(* Logix 5000 project; controller FV vendor 1 type 14 code 217 rev 31.11; software revision 31.00; part 44 of 63 *)
(* tags used below, declared in another part *)
   Dummy : BOOL;
   FV_B211 : DINT[255];   // GLYCL_SEL Glycol Pump Selectio n Words
   FV_B211_3_12_OutputBit : BOOL;
   FV_B211_3_13_OutputBit : BOOL;
   FV_B211_3_14_OutputBit : BOOL;
   fv_data_file_value_to_move : DINT;
   FV_from_data_file : DINT;
   FV_from_data_offset : DINT;
   FV_FV23C : PlantItem;   // FV23C
   FV_FV23J : PlantItem;   // FV23J
   FV_FV24C : PlantItem;   // FV24C
   FV_FV24J : PlantItem;   // FV24J
   FV_FV25C : PlantItem;   // FV25C
   FV_FV25J : PlantItem;   // FV25J
   FV_FV26C : PlantItem;   // FV26C
   FV_FV26J : PlantItem;   // FV26J
   FV_FV27C : PlantItem;   // FV27C
   FV_FV27J : PlantItem;   // FV27J
   FV_FV28C : PlantItem;   // FV28C
   FV_FV28J : PlantItem;   // FV28J
   FV_FV29C : PlantItem;   // FV29C
   FV_FV29J : PlantItem;   // FV29J
   FV_FV30C : PlantItem;   // FV30C
   FV_FV30J : PlantItem;   // FV30J
   FV_FV31C : PlantItem;   // FV31C
   FV_FV31J : PlantItem;   // FV31J
   FV_N110 : INT[255];   // FV DATA 0 CURRENT FV DATA
   FV_N111 : INT[50];   // FV1, CURRENT FV DATA
   FV_N112 : INT[50];   // FV2, CURRENT FV DATA
   FV_N113 : INT[50];   // FV3, CURRENT FV DATA
   FV_N114 : INT[50];   // FV4, CURRENT FV DATA
   FV_N115 : INT[50];   // FV5, CURRENT FV DATA
   FV_N116 : INT[50];   // FV6, CURRENT FV DATA
   FV_N117 : INT[50];   // FV7, CURRENT FV DATA
   FV_N118 : INT[50];   // FV8, CURRENT FV DATA
   FV_N119 : INT[50];   // FV9, CURRENT FV DATA
   FV_N120 : INT[50];   // FV10, CURRENT FV DATA
   FV_N121 : INT[50];   // FV11, CURRENT FV DATA
   FV_N122 : INT[50];   // FV12, CURRENT FV DATA
   FV_N123 : INT[50];   // FV13, CURRENT FV DATA
   FV_N124 : INT[50];   // FV14, CURRENT FV DATA
   FV_N125 : INT[50];   // FV15, CURRENT FV DATA
   FV_N126 : INT[50];   // FV16, CURRENT FV DATA
   FV_N127 : INT[50];   // FV17, CURRENT FV DATA
   FV_N128 : INT[50];   // FV18, CURRENT FV DATA
   FV_N129 : INT[50];   // FV19, CURRENT FV DATA
   FV_N130 : INT[50];   // FV20, CURRENT FV DATA
   FV_N131 : INT[50];   // FV21, CURRENT FV DATA
   FV_N132 : INT[50];   // FV22, CURRENT FV DATA
   FV_N133 : INT[50];   // FV23, CURRENT FV DATA
   FV_N134 : INT[50];   // FV24, CURRENT FV DATA
   FV_N135 : INT[50];   // FV25, CURRENT FV DATA
   FV_N136 : INT[50];   // YSV1, CURRENT FV DATA
   FV_N137 : INT[50];   // YSV2, CURRENT FV DATA
   FV_N138 : INT[50];   // YSV3, CURRENT FV DATA
   FV_N139 : INT[255];   // YST1
   FV_N140 : INT[255];   // YST2
   FV_N141 : INT[255];   // YSV1 DATA
   FV_N142 : INT[255];   // YSV2 DATA
   FV_N143 : INT[255];   // YSV3 DATA
   FV_N144 : INT[255];   // YST1 DATA
   FV_N145 : INT[255];   // YST2 DATA
   FV_N146 : INT[50];   // FV26, CURRENT FV DATA
   FV_N147 : INT[50];   // FV27, CURRENT FV DATA
   FV_N148 : INT[50];   // FV28, CURRENT FV DATA
   FV_N149 : INT[50];   // FV29, CURRENT FV DATA
   FV_N150 : INT[50];   // FV30, CURRENT FV DATA
   FV_N151 : INT[50];   // FV31, CURRENT FV DATA
   FV_N210 : INT[255];   // GLYCL_PTRS
   FV_PUMP1 : PlantItem;   // PUMP1
   FV_PUMP2 : PlantItem;   // PUMP2
   FV_PUMP3 : PlantItem;   // PUMP3
   FV_R6 : CONTROL[5];
   FV_SFile : INT[255];   // SLC Equivalent System File, So Original Code Can Remain
   FV_T212 : TIMER[5];
   FV_YSV1CV : PlantItem;   // YSV1CV
   FV_YSV1J : PlantItem;   // YSV1J
   FV_YSV2CV : PlantItem;   // YSV2CV
   FV_YSV2J : PlantItem;   // YSV2J
   FV_YSV3J : PlantItem;   // YSV3J
   MV_YST_Levels : REAL[2];
   YP_AV2 : PlantItem;   // AV2
   YST_BL_PMP_ON : BOOL;   // Blunger Pump
(* FV_Common, continued *)

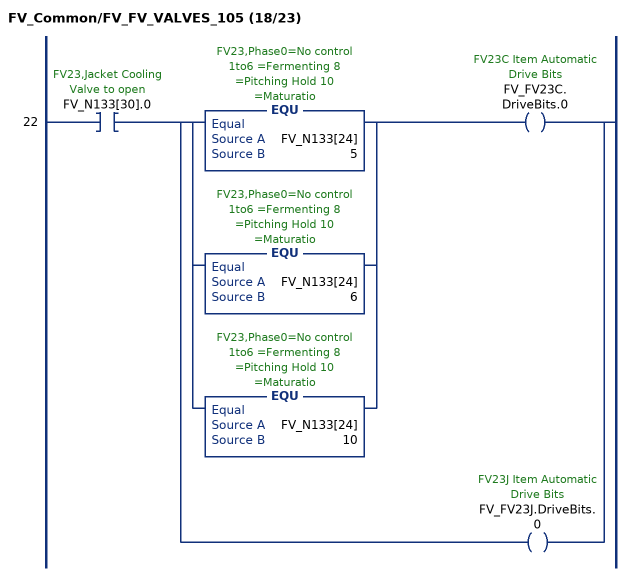
   [picture p944: FV_Common/FV_FV_VALVES_105 rungs 22-22]
   22: XIC(FV_N133[30].0)[[EQU(FV_N133[24],5) ,EQU(FV_N133[24],6) ,EQU(FV_N133[24],10) ] OTE(FV_FV23C.DriveBits.0) ,OTE(FV_FV23J.DriveBits.0) ];
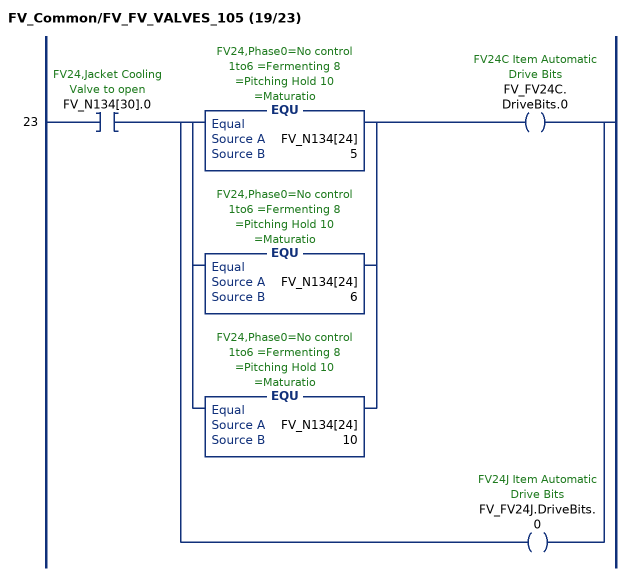
   23: XIC(FV_N134[30].0)[[EQU(FV_N134[24],5) ,EQU(FV_N134[24],6) ,EQU(FV_N134[24],10) ] OTE(FV_FV24C.DriveBits.0) ,OTE(FV_FV24J.DriveBits.0) ];
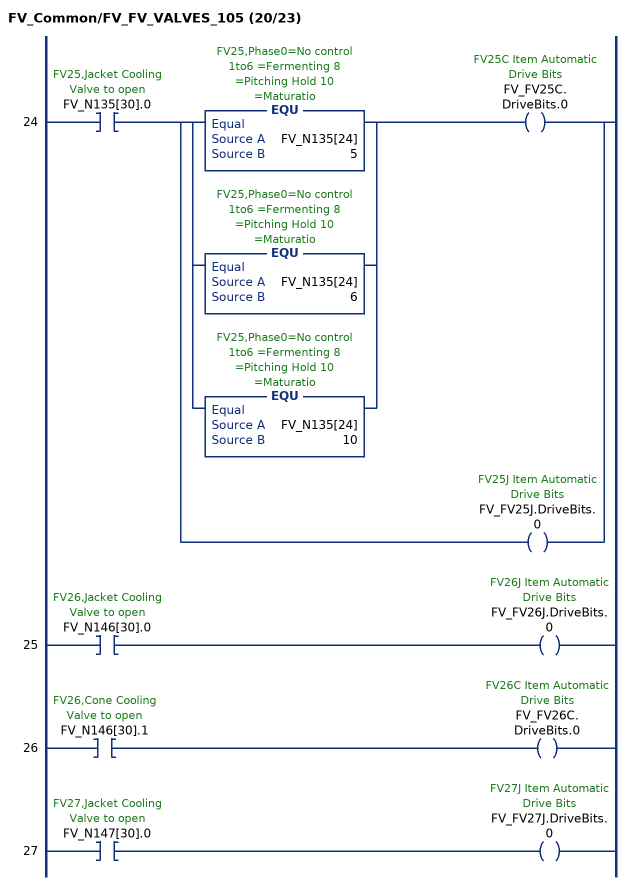
   24: XIC(FV_N135[30].0)[[EQU(FV_N135[24],5) ,EQU(FV_N135[24],6) ,EQU(FV_N135[24],10) ] OTE(FV_FV25C.DriveBits.0) ,OTE(FV_FV25J.DriveBits.0) ];
   25: XIC(FV_N146[30].0)OTE(FV_FV26J.DriveBits.0);
   26: XIC(FV_N146[30].1)OTE(FV_FV26C.DriveBits.0);
   27: XIC(FV_N147[30].0)OTE(FV_FV27J.DriveBits.0);
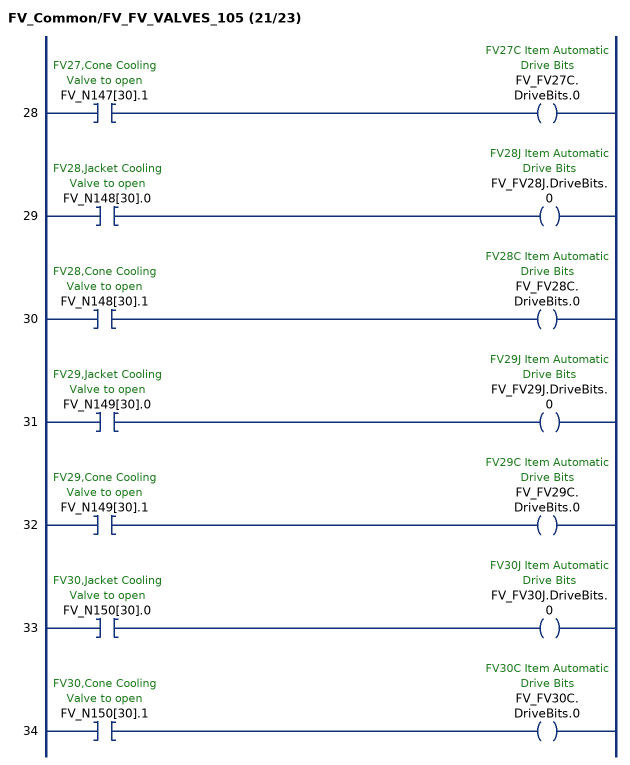
   28: XIC(FV_N147[30].1)OTE(FV_FV27C.DriveBits.0);
   29: XIC(FV_N148[30].0)OTE(FV_FV28J.DriveBits.0);
   30: XIC(FV_N148[30].1)OTE(FV_FV28C.DriveBits.0);
   31: XIC(FV_N149[30].0)OTE(FV_FV29J.DriveBits.0);
   32: XIC(FV_N149[30].1)OTE(FV_FV29C.DriveBits.0);
   33: XIC(FV_N150[30].0)OTE(FV_FV30J.DriveBits.0);
   34: XIC(FV_N150[30].1)OTE(FV_FV30C.DriveBits.0);
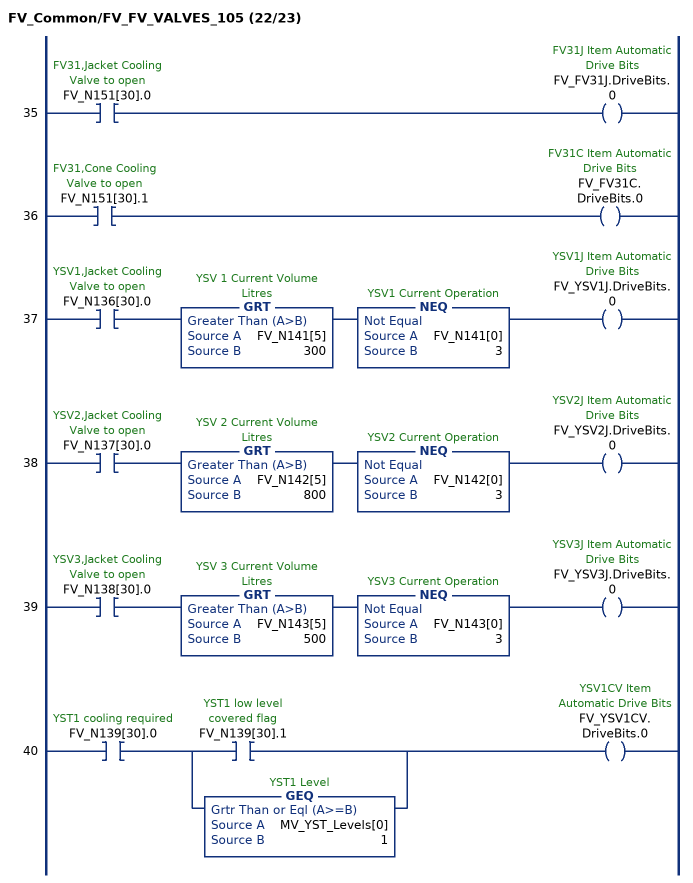
   35: XIC(FV_N151[30].0)OTE(FV_FV31J.DriveBits.0);
   36: XIC(FV_N151[30].1)OTE(FV_FV31C.DriveBits.0);
   37: XIC(FV_N136[30].0)GRT(FV_N141[5],300)NEQ(FV_N141[0],3)OTE(FV_YSV1J.DriveBits.0);
   38: XIC(FV_N137[30].0)GRT(FV_N142[5],800)NEQ(FV_N142[0],3)OTE(FV_YSV2J.DriveBits.0);
   39: XIC(FV_N138[30].0)GRT(FV_N143[5],500)NEQ(FV_N143[0],3)OTE(FV_YSV3J.DriveBits.0);
   40: XIC(FV_N139[30].0)[XIC(FV_N139[30].1) ,GEQ(MV_YST_Levels[0],1) ]OTE(FV_YSV1CV.DriveBits.0);
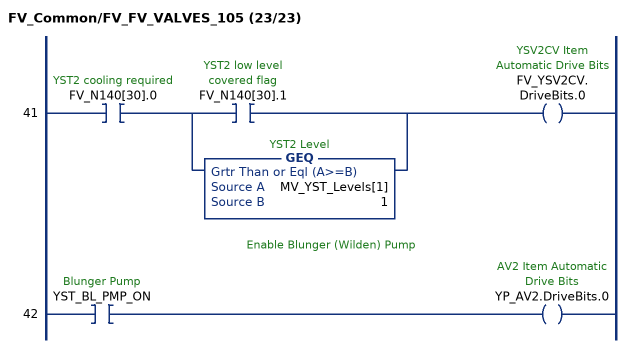
   41: XIC(FV_N140[30].0)[XIC(FV_N140[30].1) ,GEQ(MV_YST_Levels[1],1) ]OTE(FV_YSV2CV.DriveBits.0);
   // Enable Blunger (Wilden) Pump
   42: XIC(YST_BL_PMP_ON)OTE(YP_AV2.DriveBits.0);
END_ROUTINE

ROUTINE FV_Get_FV_Datafile_Value   (* ladder *)
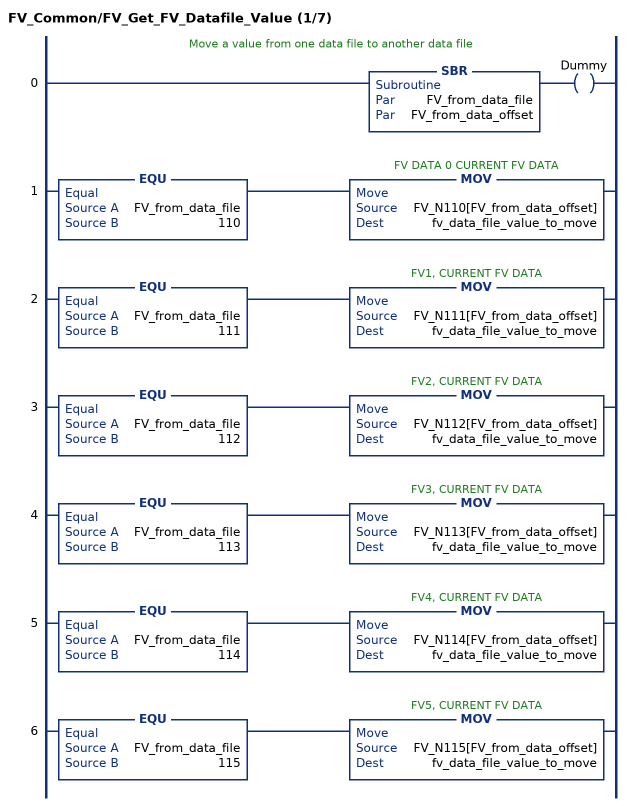
   // Move a value from one data file to another data file
   0: SBR(FV_from_data_file,FV_from_data_offset)OTE(Dummy);
   1: EQU(FV_from_data_file,110)MOV(FV_N110[FV_from_data_offset],fv_data_file_value_to_move);
   2: EQU(FV_from_data_file,111)MOV(FV_N111[FV_from_data_offset],fv_data_file_value_to_move);
   3: EQU(FV_from_data_file,112)MOV(FV_N112[FV_from_data_offset],fv_data_file_value_to_move);
   4: EQU(FV_from_data_file,113)MOV(FV_N113[FV_from_data_offset],fv_data_file_value_to_move);
   5: EQU(FV_from_data_file,114)MOV(FV_N114[FV_from_data_offset],fv_data_file_value_to_move);
   6: EQU(FV_from_data_file,115)MOV(FV_N115[FV_from_data_offset],fv_data_file_value_to_move);
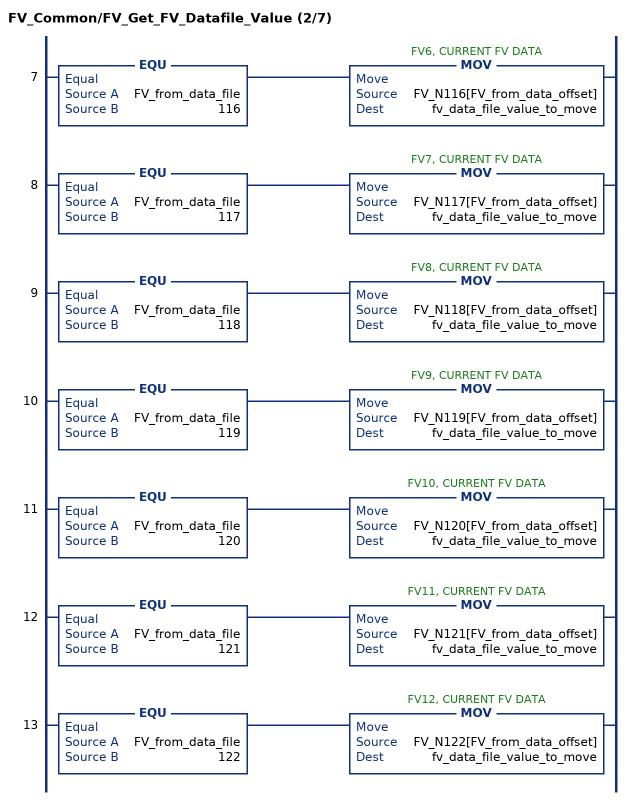
   7: EQU(FV_from_data_file,116)MOV(FV_N116[FV_from_data_offset],fv_data_file_value_to_move);
   8: EQU(FV_from_data_file,117)MOV(FV_N117[FV_from_data_offset],fv_data_file_value_to_move);
   9: EQU(FV_from_data_file,118)MOV(FV_N118[FV_from_data_offset],fv_data_file_value_to_move);
   10: EQU(FV_from_data_file,119)MOV(FV_N119[FV_from_data_offset],fv_data_file_value_to_move);
   11: EQU(FV_from_data_file,120)MOV(FV_N120[FV_from_data_offset],fv_data_file_value_to_move);
   12: EQU(FV_from_data_file,121)MOV(FV_N121[FV_from_data_offset],fv_data_file_value_to_move);
   13: EQU(FV_from_data_file,122)MOV(FV_N122[FV_from_data_offset],fv_data_file_value_to_move);
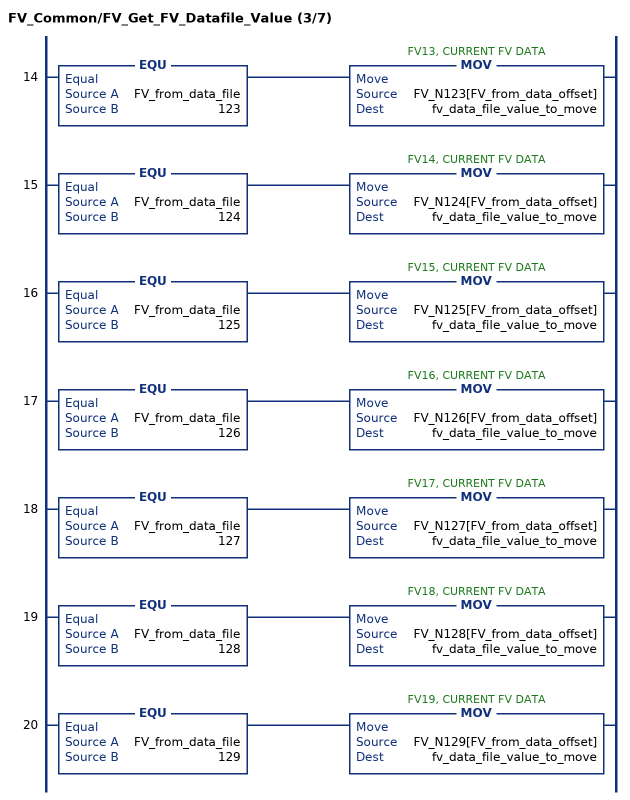
   14: EQU(FV_from_data_file,123)MOV(FV_N123[FV_from_data_offset],fv_data_file_value_to_move);
   15: EQU(FV_from_data_file,124)MOV(FV_N124[FV_from_data_offset],fv_data_file_value_to_move);
   16: EQU(FV_from_data_file,125)MOV(FV_N125[FV_from_data_offset],fv_data_file_value_to_move);
   17: EQU(FV_from_data_file,126)MOV(FV_N126[FV_from_data_offset],fv_data_file_value_to_move);
   18: EQU(FV_from_data_file,127)MOV(FV_N127[FV_from_data_offset],fv_data_file_value_to_move);
   19: EQU(FV_from_data_file,128)MOV(FV_N128[FV_from_data_offset],fv_data_file_value_to_move);
   20: EQU(FV_from_data_file,129)MOV(FV_N129[FV_from_data_offset],fv_data_file_value_to_move);
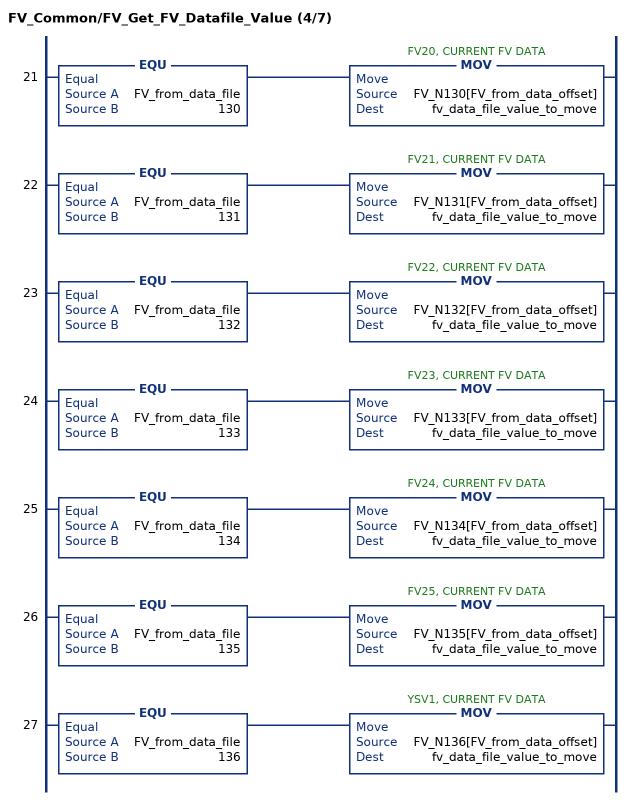
   21: EQU(FV_from_data_file,130)MOV(FV_N130[FV_from_data_offset],fv_data_file_value_to_move);
   22: EQU(FV_from_data_file,131)MOV(FV_N131[FV_from_data_offset],fv_data_file_value_to_move);
   23: EQU(FV_from_data_file,132)MOV(FV_N132[FV_from_data_offset],fv_data_file_value_to_move);
   24: EQU(FV_from_data_file,133)MOV(FV_N133[FV_from_data_offset],fv_data_file_value_to_move);
   25: EQU(FV_from_data_file,134)MOV(FV_N134[FV_from_data_offset],fv_data_file_value_to_move);
   26: EQU(FV_from_data_file,135)MOV(FV_N135[FV_from_data_offset],fv_data_file_value_to_move);
   27: EQU(FV_from_data_file,136)MOV(FV_N136[FV_from_data_offset],fv_data_file_value_to_move);
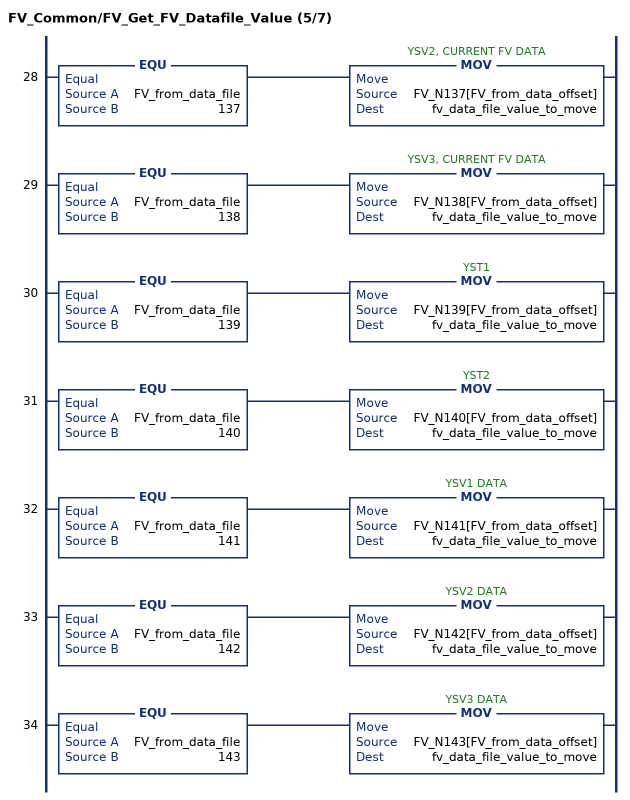
   28: EQU(FV_from_data_file,137)MOV(FV_N137[FV_from_data_offset],fv_data_file_value_to_move);
   29: EQU(FV_from_data_file,138)MOV(FV_N138[FV_from_data_offset],fv_data_file_value_to_move);
   30: EQU(FV_from_data_file,139)MOV(FV_N139[FV_from_data_offset],fv_data_file_value_to_move);
   31: EQU(FV_from_data_file,140)MOV(FV_N140[FV_from_data_offset],fv_data_file_value_to_move);
   32: EQU(FV_from_data_file,141)MOV(FV_N141[FV_from_data_offset],fv_data_file_value_to_move);
   33: EQU(FV_from_data_file,142)MOV(FV_N142[FV_from_data_offset],fv_data_file_value_to_move);
   34: EQU(FV_from_data_file,143)MOV(FV_N143[FV_from_data_offset],fv_data_file_value_to_move);
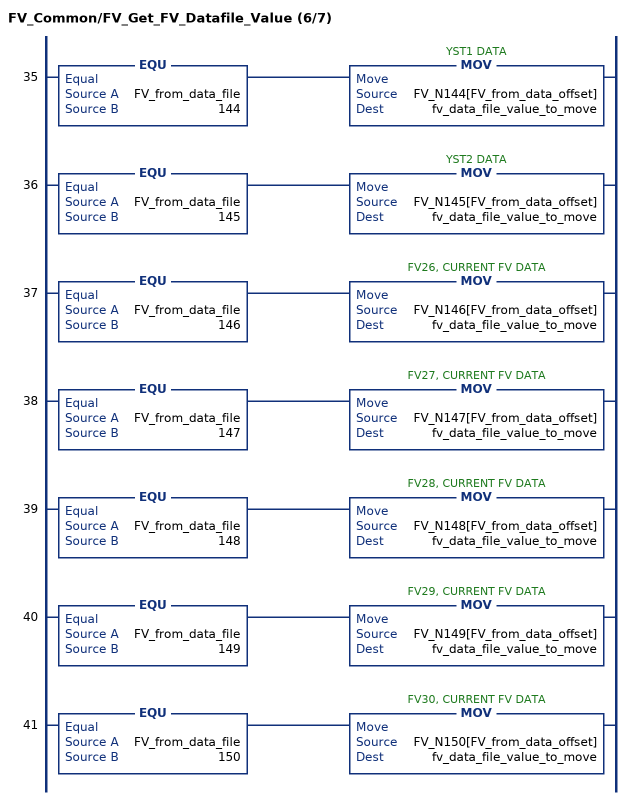
   35: EQU(FV_from_data_file,144)MOV(FV_N144[FV_from_data_offset],fv_data_file_value_to_move);
   36: EQU(FV_from_data_file,145)MOV(FV_N145[FV_from_data_offset],fv_data_file_value_to_move);
   37: EQU(FV_from_data_file,146)MOV(FV_N146[FV_from_data_offset],fv_data_file_value_to_move);
   38: EQU(FV_from_data_file,147)MOV(FV_N147[FV_from_data_offset],fv_data_file_value_to_move);
   39: EQU(FV_from_data_file,148)MOV(FV_N148[FV_from_data_offset],fv_data_file_value_to_move);
   40: EQU(FV_from_data_file,149)MOV(FV_N149[FV_from_data_offset],fv_data_file_value_to_move);
   41: EQU(FV_from_data_file,150)MOV(FV_N150[FV_from_data_offset],fv_data_file_value_to_move);
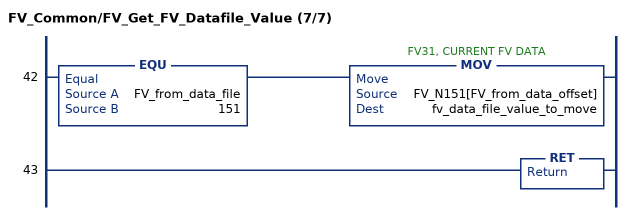
   42: EQU(FV_from_data_file,151)MOV(FV_N151[FV_from_data_offset],fv_data_file_value_to_move);
   43: RET();
END_ROUTINE

ROUTINE FV_GLYCL_PMPS_110   (* ladder *)
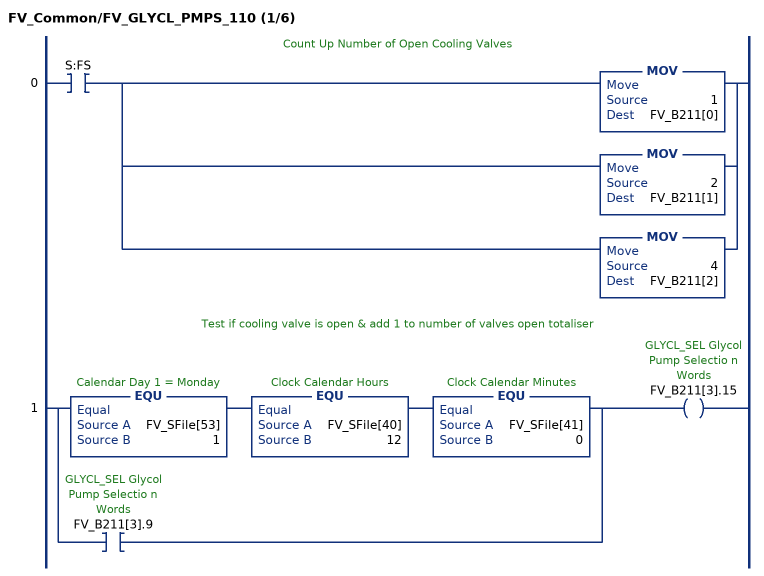
   // Count Up Number of Open Cooling Valves
   0: XIC(S:FS)[MOV(1,FV_B211[0]) ,MOV(2,FV_B211[1]) ,MOV(4,FV_B211[2]) ];
   // Test if cooling valve is open & add 1 to number of valves open totaliser
   1: [EQU(FV_SFile[53],1) EQU(FV_SFile[40],12) EQU(FV_SFile[41],0) ,XIC(FV_B211[3].9) ]OTE(FV_B211[3].15);
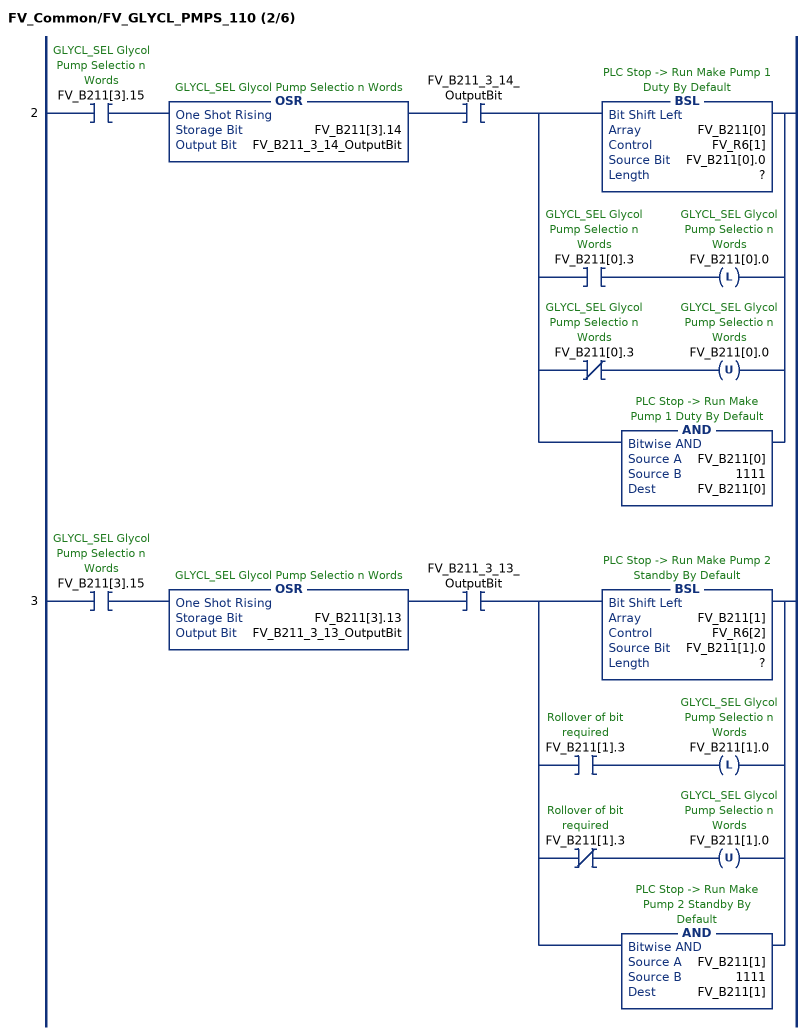
   2: XIC(FV_B211[3].15)OSR(FV_B211[3].14,FV_B211_3_14_OutputBit)XIC(FV_B211_3_14_OutputBit)[BSL(FV_B211[0],FV_R6[1],FV_B211[0].0,?) ,XIC(FV_B211[0].3) OTL(FV_B211[0].0) ,XIO(FV_B211[0].3) OTU(FV_B211[0].0) ,AND(FV_B211[0],1111,FV_B211[0]) ];
   3: XIC(FV_B211[3].15)OSR(FV_B211[3].13,FV_B211_3_13_OutputBit)XIC(FV_B211_3_13_OutputBit)[BSL(FV_B211[1],FV_R6[2],FV_B211[1].0,?) ,XIC(FV_B211[1].3) OTL(FV_B211[1].0) ,XIO(FV_B211[1].3) OTU(FV_B211[1].0) ,AND(FV_B211[1],1111,FV_B211[1]) ];
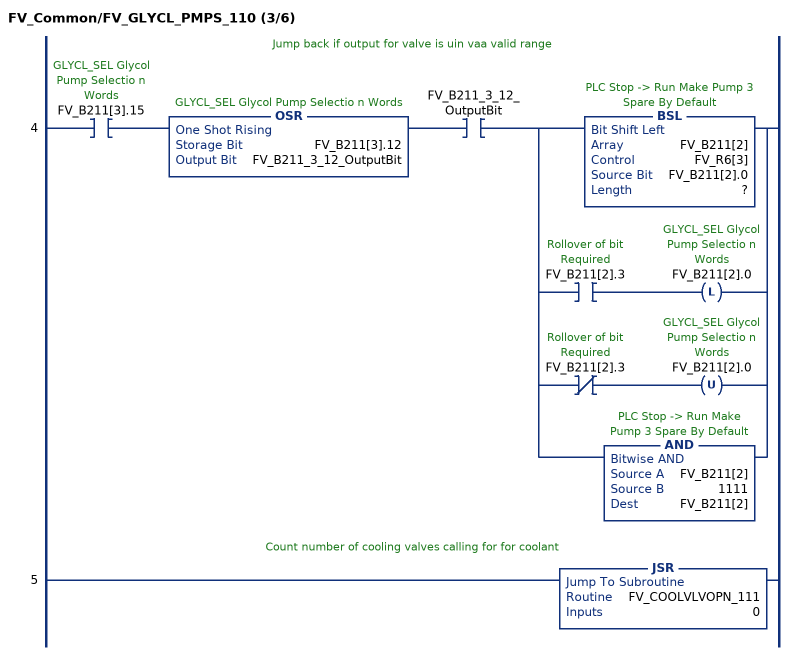
   // Jump back if output for valve is uin vaa valid range
   4: XIC(FV_B211[3].15)OSR(FV_B211[3].12,FV_B211_3_12_OutputBit)XIC(FV_B211_3_12_OutputBit)[BSL(FV_B211[2],FV_R6[3],FV_B211[2].0,?) ,XIC(FV_B211[2].3) OTL(FV_B211[2].0) ,XIO(FV_B211[2].3) OTU(FV_B211[2].0) ,AND(FV_B211[2],1111,FV_B211[2]) ];
   // Count number of cooling valves calling for for coolant
   5: JSR(FV_COOLVLVOPN_111,0);
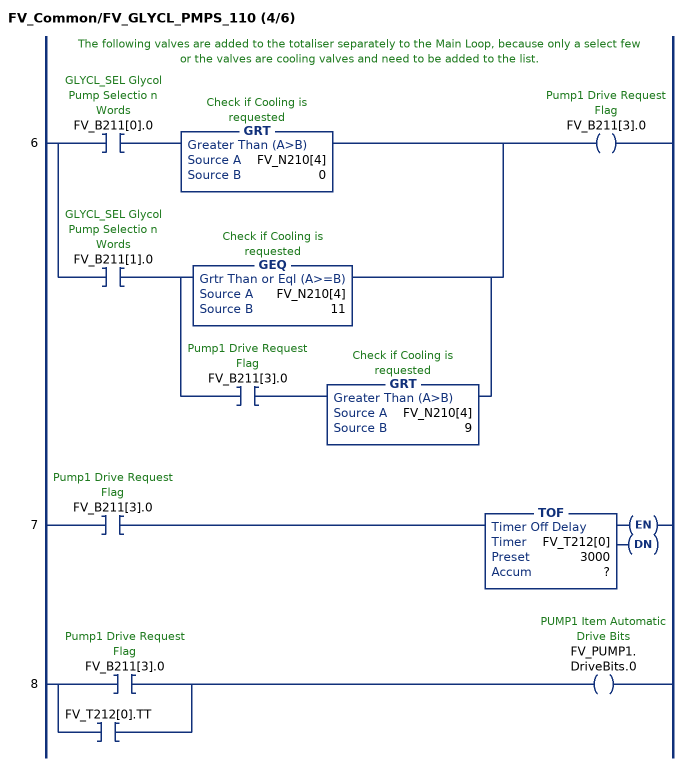
   // The following valves are added to the totaliser separately to the Main Loop, because only a select few or the valves are cooling valves and need to be added to the list.
   6: [XIC(FV_B211[0].0) GRT(FV_N210[4],0) ,XIC(FV_B211[1].0) [GEQ(FV_N210[4],11) ,XIC(FV_B211[3].0) GRT(FV_N210[4],9) ] ]OTE(FV_B211[3].0);
   7: XIC(FV_B211[3].0)TOF(FV_T212[0],?,?);
   8: [XIC(FV_B211[3].0) ,XIC(FV_T212[0].TT) ]OTE(FV_PUMP1.DriveBits.0);
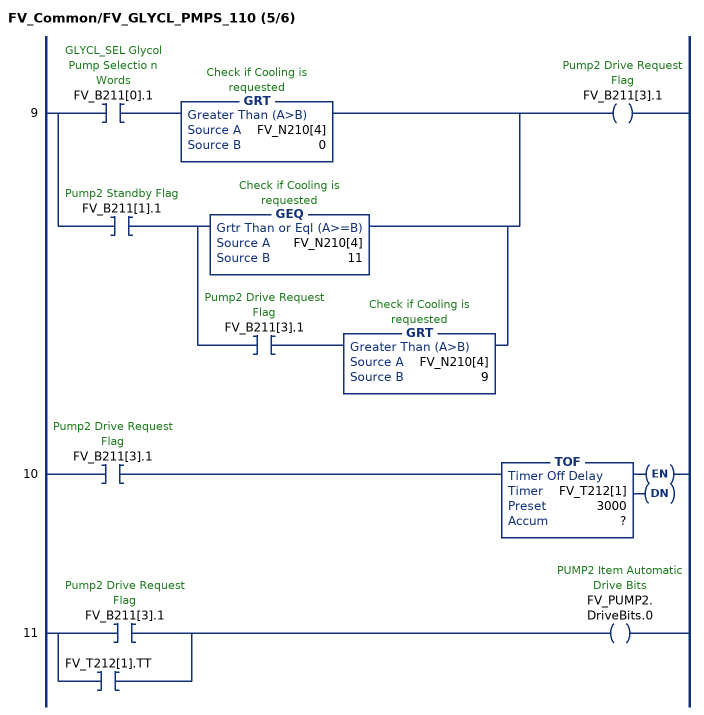
   9: [XIC(FV_B211[0].1) GRT(FV_N210[4],0) ,XIC(FV_B211[1].1) [GEQ(FV_N210[4],11) ,XIC(FV_B211[3].1) GRT(FV_N210[4],9) ] ]OTE(FV_B211[3].1);
   10: XIC(FV_B211[3].1)TOF(FV_T212[1],?,?);
   11: [XIC(FV_B211[3].1) ,XIC(FV_T212[1].TT) ]OTE(FV_PUMP2.DriveBits.0);
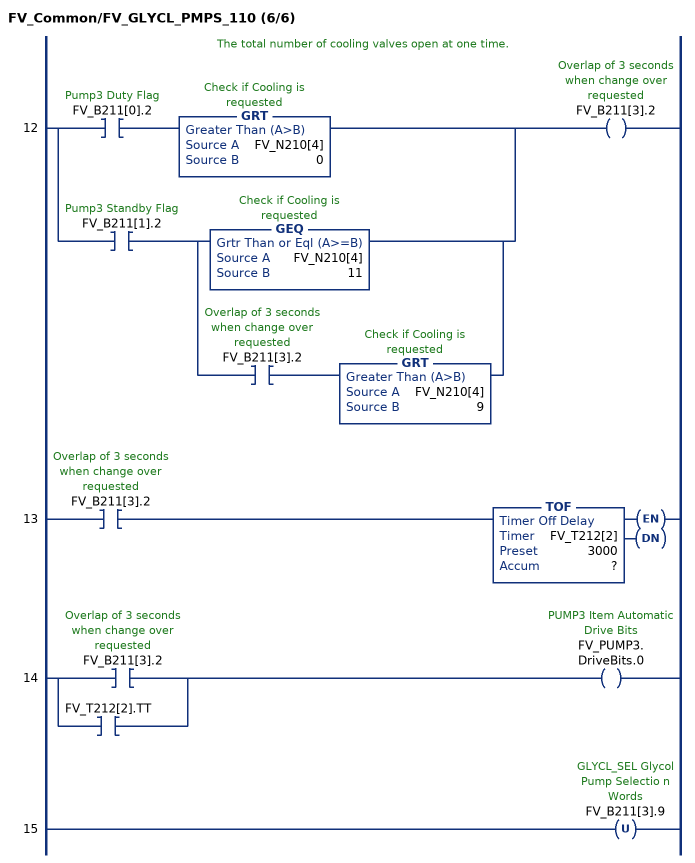
   // The total number of cooling valves open at one time.
   12: [XIC(FV_B211[0].2) GRT(FV_N210[4],0) ,XIC(FV_B211[1].2) [GEQ(FV_N210[4],11) ,XIC(FV_B211[3].2) GRT(FV_N210[4],9) ] ]OTE(FV_B211[3].2);
   13: XIC(FV_B211[3].2)TOF(FV_T212[2],?,?);
   14: [XIC(FV_B211[3].2) ,XIC(FV_T212[2].TT) ]OTE(FV_PUMP3.DriveBits.0);
   15: OTU(FV_B211[3].9);
END_ROUTINE
